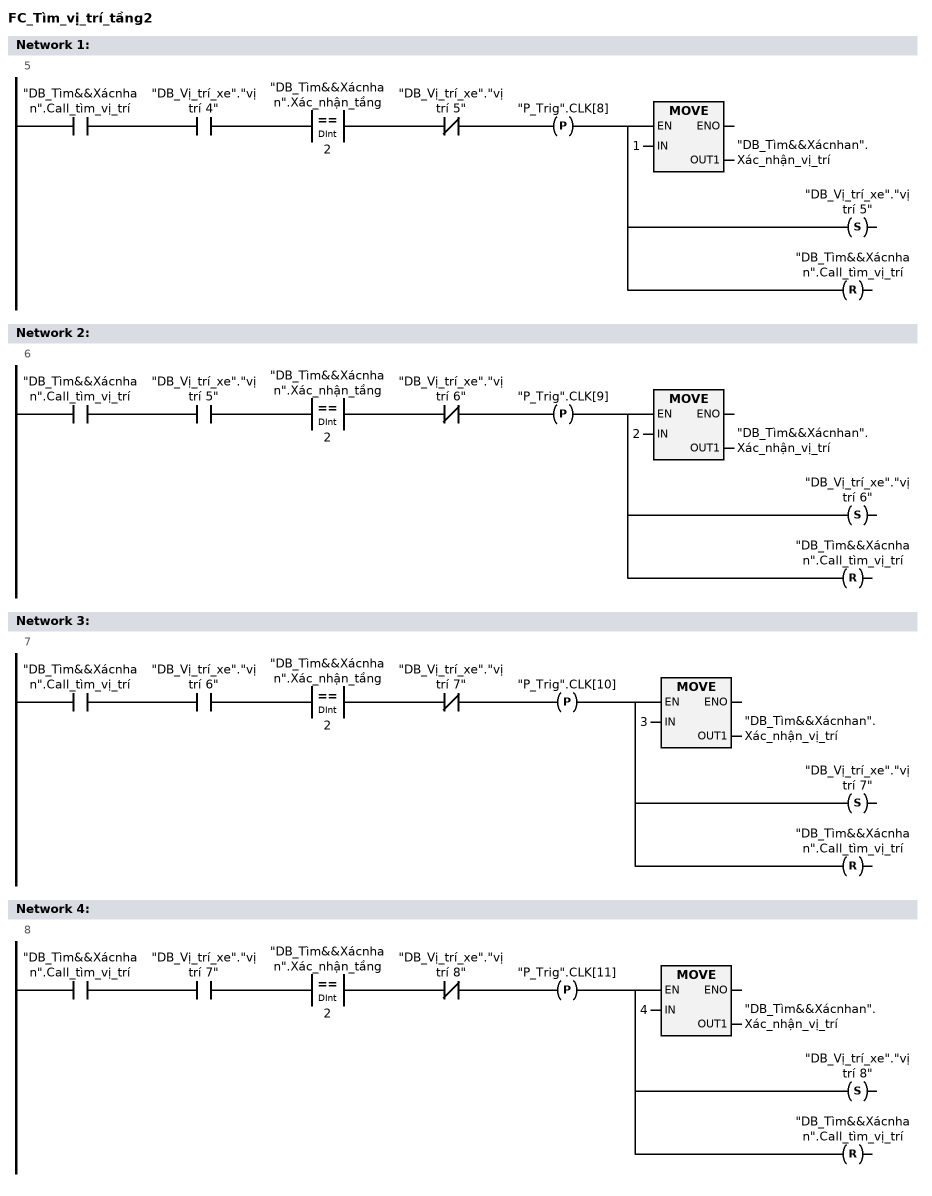
   RUNG wire#powerrail
      Contact( "DB_Tìm&&Xácnhan".Call_tìm_vị_trí )
      Contact( "DB_Vị_trí_xe"."vị trí 4" )
      { S7_Templates := "SrcType := DInt" } EQ_Contact(in1 := "DB_Tìm&&Xácnhan".Xác_nhận_tầng, in2 := 2)
      I_Contact( "DB_Vị_trí_xe"."vị trí 5" )
      P_Trig( "P_Trig".CLK[8] )
      wire#w1
      Move(in := 1, out1 => "DB_Tìm&&Xácnhan".Xác_nhận_vị_trí)
   END_RUNG
   RUNG wire#w1
      S_Coil( "DB_Vị_trí_xe"."vị trí 5" )
   END_RUNG
   RUNG wire#w1
      R_Coil( "DB_Tìm&&Xácnhan".Call_tìm_vị_trí )
   END_RUNG
   // the same network as SCL:
   #_w1 := "DB_Tìm&&Xácnhan".Call_tìm_vị_trí AND "DB_Vị_trí_xe"."vị trí 4" AND ("DB_Tìm&&Xácnhan".Xác_nhận_tầng = 2) AND NOT "DB_Vị_trí_xe"."vị trí 5";
   #_w2 := #_w1 AND NOT "P_Trig".CLK[8];   // rising edge
   "P_Trig".CLK[8] := #_w1;
   IF #_w2 THEN
       "DB_Tìm&&Xácnhan".Xác_nhận_vị_trí := 1;
       "DB_Vị_trí_xe"."vị trí 5" := TRUE;
       "DB_Tìm&&Xácnhan".Call_tìm_vị_trí := FALSE;
   END_IF;
END_REGION

REGION Network 2
   // 6
   RUNG wire#powerrail
      Contact( "DB_Tìm&&Xácnhan".Call_tìm_vị_trí )
      Contact( "DB_Vị_trí_xe"."vị trí 5" )
      { S7_Templates := "SrcType := DInt" } EQ_Contact(in1 := "DB_Tìm&&Xácnhan".Xác_nhận_tầng, in2 := 2)
      I_Contact( "DB_Vị_trí_xe"."vị trí 6" )
      P_Trig( "P_Trig".CLK[9] )
      wire#w1
      Move(in := 2, out1 => "DB_Tìm&&Xácnhan".Xác_nhận_vị_trí)
   END_RUNG
   RUNG wire#w1
      S_Coil( "DB_Vị_trí_xe"."vị trí 6" )
   END_RUNG
   RUNG wire#w1
      R_Coil( "DB_Tìm&&Xácnhan".Call_tìm_vị_trí )
   END_RUNG
   // the same network as SCL:
   #_w1 := "DB_Tìm&&Xácnhan".Call_tìm_vị_trí AND "DB_Vị_trí_xe"."vị trí 5" AND ("DB_Tìm&&Xácnhan".Xác_nhận_tầng = 2) AND NOT "DB_Vị_trí_xe"."vị trí 6";
   #_w2 := #_w1 AND NOT "P_Trig".CLK[9];   // rising edge
   "P_Trig".CLK[9] := #_w1;
   IF #_w2 THEN
       "DB_Tìm&&Xácnhan".Xác_nhận_vị_trí := 2;
       "DB_Vị_trí_xe"."vị trí 6" := TRUE;
       "DB_Tìm&&Xácnhan".Call_tìm_vị_trí := FALSE;
   END_IF;
END_REGION

REGION Network 3
   // 7
   RUNG wire#powerrail
      Contact( "DB_Tìm&&Xácnhan".Call_tìm_vị_trí )
      Contact( "DB_Vị_trí_xe"."vị trí 6" )
      { S7_Templates := "SrcType := DInt" } EQ_Contact(in1 := "DB_Tìm&&Xácnhan".Xác_nhận_tầng, in2 := 2)
      I_Contact( "DB_Vị_trí_xe"."vị trí 7" )
      P_Trig( "P_Trig".CLK[10] )
      wire#w1
      Move(in := 3, out1 => "DB_Tìm&&Xácnhan".Xác_nhận_vị_trí)
   END_RUNG
   RUNG wire#w1
      S_Coil( "DB_Vị_trí_xe"."vị trí 7" )
   END_RUNG
   RUNG wire#w1
      R_Coil( "DB_Tìm&&Xácnhan".Call_tìm_vị_trí )
   END_RUNG
   // the same network as SCL:
   #_w1 := "DB_Tìm&&Xácnhan".Call_tìm_vị_trí AND "DB_Vị_trí_xe"."vị trí 6" AND ("DB_Tìm&&Xácnhan".Xác_nhận_tầng = 2) AND NOT "DB_Vị_trí_xe"."vị trí 7";
   #_w2 := #_w1 AND NOT "P_Trig".CLK[10];   // rising edge
   "P_Trig".CLK[10] := #_w1;
   IF #_w2 THEN
       "DB_Tìm&&Xácnhan".Xác_nhận_vị_trí := 3;
       "DB_Vị_trí_xe"."vị trí 7" := TRUE;
       "DB_Tìm&&Xácnhan".Call_tìm_vị_trí := FALSE;
   END_IF;
END_REGION

REGION Network 4
   // 8
   RUNG wire#powerrail
      Contact( "DB_Tìm&&Xácnhan".Call_tìm_vị_trí )
      Contact( "DB_Vị_trí_xe"."vị trí 7" )
      { S7_Templates := "SrcType := DInt" } EQ_Contact(in1 := "DB_Tìm&&Xácnhan".Xác_nhận_tầng, in2 := 2)
      I_Contact( "DB_Vị_trí_xe"."vị trí 8" )
      P_Trig( "P_Trig".CLK[11] )
      wire#w1
      Move(in := 4, out1 => "DB_Tìm&&Xácnhan".Xác_nhận_vị_trí)
   END_RUNG
   RUNG wire#w1
      S_Coil( "DB_Vị_trí_xe"."vị trí 8" )
   END_RUNG
   RUNG wire#w1
      R_Coil( "DB_Tìm&&Xácnhan".Call_tìm_vị_trí )
   END_RUNG
   // the same network as SCL:
   #_w1 := "DB_Tìm&&Xácnhan".Call_tìm_vị_trí AND "DB_Vị_trí_xe"."vị trí 7" AND ("DB_Tìm&&Xácnhan".Xác_nhận_tầng = 2) AND NOT "DB_Vị_trí_xe"."vị trí 8";
   #_w2 := #_w1 AND NOT "P_Trig".CLK[11];   // rising edge
   "P_Trig".CLK[11] := #_w1;
   IF #_w2 THEN
       "DB_Tìm&&Xácnhan".Xác_nhận_vị_trí := 4;
       "DB_Vị_trí_xe"."vị trí 8" := TRUE;
       "DB_Tìm&&Xácnhan".Call_tìm_vị_trí := FALSE;
   END_IF;
END_REGION
END_FUNCTION

FUNCTION "FC_tìm_vị_trí" : Void   // FC8, LAD
{ S7_Optimized_Access := 'TRUE' }
VERSION : 0.1
BEGIN

REGION Network 1
   // Tìm trong tầng , coi vị trí trống,move hướng(1-4),đánh dấu vị trí,kết thuc gọi tìm vị trí
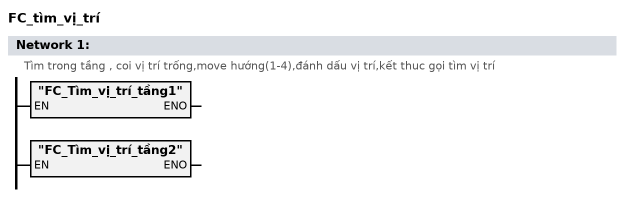
   RUNG wire#powerrail
      "FC_Tìm_vị_trí_tầng1"()
   END_RUNG
   RUNG wire#powerrail
      "FC_Tìm_vị_trí_tầng2"()
   END_RUNG
   // the same network as SCL:
   "FC_Tìm_vị_trí_tầng1"();
   "FC_Tìm_vị_trí_tầng2"();
END_REGION
END_FUNCTION

(* ===== HMI "HMI_RT_1" =====
connection "HMI_Connection_1": ETHERNET, ILRT_S7_1500_OMS

HMI tags "Default tag table"
   "DB_AxisPanel_Lift_Job_Velocity" : Real = PLC DB_AxisPanel.Lift.Job.Velocity, T1s

HMI tags "Operater"
   "DB_Operater_Confirm_Gửi" : Bool = PLC DB_Operater.Confirm_Gửi AT %DB6.DBX0.0, T100ms
   "DB_Operater_Confirm_Lấy" : Bool = PLC DB_Operater.Confirm_Lấy AT %DB6.DBX0.1, T100ms
   "DB_Operater_Scada_Gửi_Xe" : Bool = PLC DB_Operater.Scada_Gửi_Xe AT %DB6.DBX0.3, T100ms
   "DB_Operater_Scada_Lấy_Xe" : Bool = PLC DB_Operater.Scada_Lấy_Xe AT %DB6.DBX0.4, T100ms
   "DB_Operater_ConfirmRFID" : Bool = PLC DB_Operater.ConfirmRFID AT %DB6.DBX0.2, T100ms
   "DB_Operater_Scada_Home_Lift" : Bool = PLC DB_Operater.Scada_Home_Lift AT %DB6.DBX0.6, T100ms
   "DB_Operater_AutoMan" : Bool = PLC DB_Operater.Auto/Man AT %DB6.DBX1.0, T100ms
   "DB_Operater_Static_Mode" : Int = PLC DB_Operater.Static_Mode AT %DB6.DBW2, T100ms

HMI tags "Step"
   "DB_Step_Power" : Bool = PLC DB_Step.Power, T100ms
   "DB_Step_Home_Lift" : Bool = PLC DB_Step.Home.Lift, T100ms
   "DB_Step_Home_Rotation" : Bool = PLC DB_Step.Home.Rotation, T100ms
   "DB_Step_Home_Reach" : Bool = PLC DB_Step.Home.Reach, T100ms
   "DB_Step_HomeAll" : Bool = PLC DB_Step.HomeAll, T100ms
   "DB_Step_ErorrHomeCode_Lift" : Word = PLC DB_Step.ErorrHomeCode.Lift, T100ms
   "DB_Step_ErorrHomeCode_Rotation" : Word = PLC DB_Step.ErorrHomeCode.Rotation, T100ms
   "DB_Step_ErorrHomeCode_Reach" : Word = PLC DB_Step.ErorrHomeCode.Reach, T100ms
   "DB_Step_ErrorHome_Lift" : Bool = PLC DB_Step.ErrorHome.Lift, T100ms
   "DB_Step_ErrorHome_Rotation" : Bool = PLC DB_Step.ErrorHome.Rotation, T100ms
   "DB_Step_ErrorHome_Reach" : Bool = PLC DB_Step.ErrorHome.Reach, T100ms
   "DB_Step_ErorrAbsoluteCode_Rotation" : Word = PLC DB_Step.ErorrAbsoluteCode.Rotation, T100ms
   "DB_Step_ErorrAbsoluteCode_Lift" : Word = PLC DB_Step.ErorrAbsoluteCode.Lift, T100ms
   "DB_Step_ErorrAbsoluteCode_Reach" : Word = PLC DB_Step.ErorrAbsoluteCode.Reach, T100ms
   "DB_Step_ErrorAbsolute_Lift" : Bool = PLC DB_Step.ErrorAbsolute.Lift, T100ms
   "DB_Step_ErrorAbsolute_Rotation" : Bool = PLC DB_Step.ErrorAbsolute.Rotation, T100ms
   "DB_Step_ErrorAbsolute_Reach" : Bool = PLC DB_Step.ErrorAbsolute.Reach, T100ms
   "DB_Step_ErrorJog_Lift" : Word = PLC DB_Step.ErrorJog.Lift, T100ms
   "DB_Step_ErrorJog_Rotation" : Word = PLC DB_Step.ErrorJog.Rotation, T100ms
   "DB_Step_ErrorJog_Reach" : Word = PLC DB_Step.ErrorJog.Reach, T100ms
   "DB_Step_Reset" : Bool = PLC DB_Step.Reset, T100ms
   "DB_Step_PowerStarted" : Bool = PLC DB_Step.PowerStarted, T100ms
   "DB_Step_HomeStarted" : Bool = PLC DB_Step.HomeStarted, T100ms
   "DB_Step_DoneHome" : Bool = PLC DB_Step.DoneHome, T100ms

HMI tags "Convert"
   "DB_Convert_Python_Floor" : Int = PLC DB_Convert.Python.Floor AT %DB14.DBW0, T1s
   "DB_Convert_Python_Location" : Int = PLC DB_Convert.Python.Location AT %DB14.DBW2, T1s
   "DB_Convert_Python_Passcodeplc" : Int = PLC DB_Convert.Python.Passcodeplc AT %DB14.DBW4, T1s
   "DB_Convert_Python_UID" : Array [0..11] of String[14] = PLC DB_Convert.Python.UID AT %DB14.DBX6.0, T1s
   "DB_Convert_Python_Receive" : String[14] = PLC DB_Convert.Python.Receive AT %DB14.DBX198.0, T1s
   "DB_Convert_Floor_Dic1" : Int = PLC DB_Convert.Floor_Dic1 AT %DB14.DBW214, T1s
   "DB_Convert_Floor_Dic2" : Int = PLC DB_Convert.Floor_Dic2 AT %DB14.DBW216, T1s
   "DB_Convert_Location" : Int = PLC DB_Convert.Location AT %DB14.DBW218, T1s
   "DB_Convert_Down" : Int = PLC DB_Convert.Down AT %DB14.DBW220, T1s
   "DB_Convert_Up" : Int = PLC DB_Convert.Up AT %DB14.DBW222, T1s
   "DB_Convert_Started" : Bool = PLC DB_Convert.Started AT %DB14.DBX224.0, T1s

HMI tags "Axis_Panel"
   "DB_AxisPanel_Lift" : UDT = PLC DB_AxisPanel.Lift, T100ms
   "DB_AxisPanel_Rotation" : UDT = PLC DB_AxisPanel.Rotation, T100ms
   "DB_AxisPanel_Reach" : UDT = PLC DB_AxisPanel.Reach, T100ms

HMI tags "Vị trí xe"
   "DB_Vị_trí_xe_vị trí 1" : Bool = PLC DB_Vị_trí_xe."vị trí 1" AT %DB2.DBX0.0, T100ms
   "DB_Vị_trí_xe_vị trí 2" : Bool = PLC DB_Vị_trí_xe."vị trí 2" AT %DB2.DBX0.1, T100ms
   "DB_Vị_trí_xe_vị trí 3" : Bool = PLC DB_Vị_trí_xe."vị trí 3" AT %DB2.DBX0.2, T100ms
   "DB_Vị_trí_xe_vị trí 4" : Bool = PLC DB_Vị_trí_xe."vị trí 4" AT %DB2.DBX0.3, T100ms
   "DB_Vị_trí_xe_vị trí 5" : Bool = PLC DB_Vị_trí_xe."vị trí 5" AT %DB2.DBX0.4, T100ms
   "DB_Vị_trí_xe_vị trí 6" : Bool = PLC DB_Vị_trí_xe."vị trí 6" AT %DB2.DBX0.5, T100ms
   "DB_Vị_trí_xe_vị trí 7" : Bool = PLC DB_Vị_trí_xe."vị trí 7" AT %DB2.DBX0.6, T100ms
   "DB_Vị_trí_xe_vị trí 8" : Bool = PLC DB_Vị_trí_xe."vị trí 8" AT %DB2.DBX0.7, T100ms
   "DB_Vị_trí_xe_tầng_1" : Bool = PLC DB_Vị_trí_xe.tầng_1 AT %DB2.DBX1.0, T100ms
   "DB_Vị_trí_xe_tầng_2" : Bool = PLC DB_Vị_trí_xe.tầng_2 AT %DB2.DBX1.1, T100ms

text list "SystemTextList_ConfigErrorAlarmTextLibrary_1": 1 'NameService configuration error: Implicit deletion. Subelement instance @6%s@ must be deleted explicitly.'; 2 'NameService configuration error: Implicit deletion. Alias/Format/Unit instance @6%s@ must be deleted explicitly.'

text list "SystemTextList_ConfigErrorAlarmTextLibrary_2": 1 'EvDpManager::cleanupDeletedDatapoint - alert handler config is deleted implicitly for deleted datapoint, @3%s@'; 2 'EvDpManager::cleanupDeletedDatapoint - alert handler config is deleted implicitly but still has overrides, @3%s@'; 3 'EvDpManager::cleanupDeletedDatapoint - default value config is deleted implicitly for deleted datapoint, @3%s@'; 4 'EvDpManager::cleanupDeletedDatapoint - default value config is deleted implicitly but still has overrides, @3%s@'; 5 'EvDpManager::cleanupDeletedDatapoint - initial value config is deleted implicitly for deleted datapoint, @3%s@'; 6 'EvDpManager::cleanupDeletedDatapoint - initial value config is deleted implicitly but still has overrides, @3%s@'; 7 'EvDpManager::cleanupDeletedDatapoint - distribution config is deleted implicitly for deleted datapoint, @3%s@'; 8 'EvDpManager::cleanupDeletedDatapoint - distribution config is deleted implicitly but still has overrides, @3%s@'; 9 'EvDpManager::cleanupDeletedDatapoint - rangeCheck config is deleted implicitly for deleted datapoint, @3%s@'; 10 'EvDpManager::cleanupDeletedDatapoint - rangeCheck config is deleted implicitly but still has overrides, @3%s@'

text list "SystemTextList_ConfigErrorAlarmTextLibrary_3": 1 'The configured data point type was deleted, but a configured type is still defined for the node type: @3%s@.'; 2 'The configured data point node type was deleted in the data point type, but a configured type is still defined for the element: @3%s@.'

text list "SystemTextList_ConfigErrorAlarmTextLibrary_4": 2 'Cycles: @6%s@ does not exist'; 3 'Alarms: @6%s@ exists already'; 4 'Tags: Address @6%s@ was rejected'; 1 'Connections: @6%s@ does not exist'; 5 'Tags: Acquisition mode @6%s@ is not supported.'; 6 'Cycles: @6%s@ was deleted but associated tags exist.'; 7 'Connections: @6%s@ was deleted but associated tags exist.'; 8 'Tags: Tag @6%s@ was rejected.'; 9 'Tags: Tag @6%s@ has an invalid value.'; 0 'Connections: Connection to @6%s@ could not be established.'; 65638 'Connections: Connection to @6%s@ could not be established.'; 65639 'Connections: @6%s@ disconnected.'; 65640 'Connections: Connection to the HMI device @6%s@ is lost.'; 65641 'Connections: Connection to the PLC @6%s@ is lost.'; 65541 'Connections: Timeout while establishing the connection to @6%s@.'; 65542 'Connections: @6%s@ faulty.'; 65543 'Connections: Connection to the HMI device disconnected. Connection @5%s@ was changed.'; 65544 'Connections: Connection to the HMI device disconnected. Driver property was changed for connection @5%s@.'

text list "SystemTextList_ConfigErrorAlarmTextLibrary_5": 1 'Connections: Lifecycle monitoring cycle must be shorter than the response time.'; 2 'Connections: Cyclic services are configured but not supported by the target device.'; 3 'Connections: Change-controlled reading is configured but not supported by the target device.'; 4 'Tags: The address @6%s@ does not exist in the PLC.'; 5 'Tags: The default conversion type for the address @6%s@ could not be determined.'; 6 'Tags: Invalid conversion type'; 7 'Cycles: Invalid conversion type. Conversion is not supported at HmiCycle.'; 4096 'Connections: Version of the address @6%s@ is not supported.'; 4097 'Connections: PROFIBUS address is not supported.'; 4098 'Connections: Softbus address is not supported.'; 4099 'Connections: Address type @6%s@ is not supported.'; 4100 'Connections: Invalid connection name @6%s@. Access point is being ignored.'; 4101 'Connections: Routing is not supported. @6%s@ is not used.'; 4102 'Connections: Routing is not supported. @6%s@ is not used.'; 4103 'Connections: Invalid IP address @6%s@'; 4104 'Connections: Invalid Named Connection @6%s@. Valid format: >VMD</>connection<'; 4105 'Connections: Invalid Named Connection @6%s@. VMD connection name is too long. Only 24 characters are permitted.'; 4106 'Connections: Invalid Named Connection @6%s@. Connection name is too long. Only 32 characters are permitted.'; 4107 'Connections: Rack number @6%s@ is outside of the permitted range (0..7)'; 4108 'Connections: Invalid Named Connection @6%s@. Rack is ignored.'; 4109 'Connections: Slot number @6%s@ is outside of the permitted range (1..32)'; 4110 'Connections: Invalid Named Connection @6%s@. Slot is ignored.'; 4111 'Connection could not be established. Maximum number of available connections (@6%s@) has been exceeded.'; 4112 'Connection aborted. No sign of life in the last @4%s@ ms.'; 4113 'Connection could not be established - @4%s@'; 4114 'Connection could not be established. The address @6%s@ cannot be used.'; 4115 'Connection could not be established. Invalid address @6%s@'; 4116 'Connection could not be established - @4%s@'

text list "SystemTextList_ConfigErrorAlarmTextLibrary_6": 1 'Connection could not be established. Application instance certificate is not configured.'; 2 'Connection could not be established. Server has rejected the client certificate. OPC UA status code @4%s@.'; 3 'Connection could not be established. Internal problem in the certificate store. OPC UA status code @4%s@'; 4 'Connection could not be established. Application instance certificate could not be loaded. OPC UA status code @4%s@'; 5 'Connection could not be established. Server has not provided a certificate. @4%s@'; 6 'Connection could not be established. Validation of server certificate has failed. OPC UA status code @4%s@.'; 7 'Connection was closed. Error during alarm synchronization. OPC UA status code @4%s@.'; 8 'Connection was closed. Alarm/event subscription has failed. The number of operations on the server has been exceeded.'; 9 'Connection was closed. Alarm/event subscription has failed. The number of alarm/event subscriptions on the server has been exceeded.'; 10 'Connection could not be established. Server reports a license problem. OPC UA status code @4%s@.'; 11 'Connection could not be established. Maximum number of server sessions has been exceeded.'; 12 'Connection could not be established. Safety configuration is inconsistent. @4%s@'; 13 'Connection could not be established. The address @4%s@ cannot be used.'; 14 'Connection could not be established. OPC UA status code @4%s@'; 15 'Connection aborted. OPC UA server was stopped.'; 16 'Connection aborted. No sign of life in the last @4%s@ ms.'; 17 'Connection was closed. OPC UA server maintenance.'; 18 'Connection could not be established. Invalid configuration of the authentication mode - @4%s@'; 19 'Connection could not be established. User could not be authenticated. OPC UA status code @4%s@'; 20 'Connection could not be established. Server does not permit anonymous connection. OPC UA status code @4%s@'; 21 'Connection could not be established. Certificate problem: Error when writing the safety-relevant data to @4%s@.'; 22 'Connection could not be established. Certificate problem: Unexpected file in the folder @4%s@ cannot be removed.'; 23 'Connection could not be established. User could not be authenticated. No user or password configured.'; 24 'Connection could not be established. Unexpected length of the server certificate. @4%s@'; 25 'Connection could not be established. @4%s@ is empty.'; 26 'Connection could not be established. @4%s@ has an unexpected format.'; 27 'Connection could not be established. Server endpoints cannot be read. OPC UA status code @4%s@'; 28 'Connection could not be established. No server endpoints were found. @4%s@'; 29 'Connection could not be established. Application instance certificate could not be found.'; 30 'Connection could not be established. Unexpected format of the certificate @4%s@.'; 31 'Connection could not be established. Unexpected format of the certificate block list @4%s@.'; 32 'Connection could not be established. User could not be authenticated. An encryption detail is invalid. @4%s@'; 34 'Connection could not be established. - The configured non-transparent redundancy mode @4%s@ is not supported.'; 101 'Tags: Address @6%s@ does not exist on the server.'; 103 'Tags: Address @6%s@ cannot be accessed.'; 104 'Tags: Acquisition mode is not supported for address @6%s@.'; 201 'Alarms: Address @6%s@ does not exist on the server.'; 202 'Alarms: Address @6%s@ cannot be used. The specified range filter is not an OPC UA Event Notifier.'; 203 'Alarms: Address @6%s@ cannot be used. The specified range filter does not exist on the server.'; 204 'Alarms: Address @6%s@ cannot be used because it is not an OPC UA event type.'; 205 'Alarms: Address @6%s@ cannot be used because the OPC UA condition type is not supported.'; 206 'Alarms: Address @6%s@ cannot be used because the event type does not exist on the server.'; 207 'Alarms: Acquisition type cannot be used for address @6%s@.'; 301 'Address @6%s@ cannot be used because the version number is missing.'; 302 'Address @6%s@ cannot be used because the version number is invalid.'; 303 'Address @6%s@ cannot be used because the number of '$' delimiters is invalid.'; 304 'Address @6%s@ cannot be used because the address type is invalid.'; 305 'Unsupported version @6%s@ of the address'; 401 'Unexpected OPC UA server response: @6%s@'

text list "SystemTextList_ConfigErrorAlarmTextLibrary_7": 1 'Messages: Invalid condition string for the alarm view @6%s@.'; 2 'Messages: Invalid status tag and bit for the alarm view @6%s@.'; 3 'Messages: Invalid control tag and bit for the alarm view @6%s@.'

text list "SystemTextList_ConfigErrorAlarmTextLibrary_8": 1 'Logs: Implicit deletion. Logging tag instance @6%s@ should be deleted but there are overloaded elements.'

text list "SystemTextList_ConfigErrorAlarmTextLibrary_9": 1 ''; 2 'Restart of the runtime is required.'; 3 'The correct storage medium must be ejected and inserted again.'

text list "SystemTextList_ConfigErrorAlarmTextLibrary_10": 1 'CDS cache - Cache folder cannot be created or reached: @6%s@'; 2 'LOC cache - Cache folder cannot be created or reached: @6%s@'

text list "SystemTextList_RuntimeCollaborationFailureReason_1": 0 'Unknown error (@3%s@)'; 1 'The system is not running or there is a network problem'; 2 'Runtime is not started on the target device.'; 3 'The System ID does not match the expected System ID (@3%s@)'; 4 'The Collaboration name does not match the expected Collaboration name '@3%s@''; 5 'Wrong or unknown certificate'; 6 'Revoked certificate'; 7 'The time difference is too big.'; 8 'No common supported message version'; 9 'System ID (@3%s@) already exists'; 10 'System name (@3%s@) already exists'; 11 'ID/Name in local configuration for Runtime Collaboration already exists'

text list "SystemTextList_S7PlusAlarmTextListCollection_1": 4096 'Connections: Connection to the PLC @4%s@ is lost'; 4097 'Connections: Connection to the HMI device @4%s@ is lost'; 4098 'Connections: Maximum number of connections exceeded - @4%s@'; 4099 'Out of resources on PLC - @4%s@'; 4100 'Legitimation failed, invalid or missing password - @4%s@'; 4101 'Request to open the connection failed - @4%s@'; 4102 'Connections: Cannot connect to PLC - @4%s@'; 4103 'Request to open the connection could not be sent'; 4104 'General certificate error for PLC - @4%s@'; 4105 'PLC certificate expired for PLC - @4%s@'; 4106 'PLC certificate is revoked for PLC - @4%s@'; 4107 'PLC certificate is untrustworthy. Manual trust is possible for - @4%s@'; 4108 'PLC certificate is untrustworthy. Manual trust is not possible for - @4%s@'

text list "SystemTextList_AllenBradleyEIPAlarmTextListCollection_7": 4096 'Connection lost on PLC side - @5%s@'; 4097 'Connection lost on HMI side - @5%s@'; 4098 'Maximum number of connections exceeded - @5%s@'; 4099 'Out of resources on PLC - @5%s@'; 4100 'Legitimation failed, invalid or missing password - @5%s@'; 4101 'Open request failed - @5%s@'; 4102 'Cannot connect to PLC - @5%s@'; 4103 'Open request could not be sent'; 4104 'root certificate expired for - @5%s@'; 4105 'PLC certificate untrusted for - @5%s@'

text list "SystemTextList_OmronEIPAlarmTextListCollection_6": 4096 'Connection lost on PLC side - @5%s@'; 4097 'Connection lost on HMI side - @5%s@'; 4098 'Maximum number of connections exceeded - @5%s@'; 4099 'Out of resources on PLC - @5%s@'; 4100 'Legitimation failed, invalid or missing password - @5%s@'; 4101 'Open request failed - @5%s@'; 4102 'Cannot connect to PLC - @5%s@'; 4103 'Open request could not be sent'; 4104 'root certificate expired for - @5%s@'; 4105 'PLC certificate untrusted for - @5%s@'

text list "SystemTextList_StdModbusTCPAlarmTextListCollection_5": 4096 'Connections: Connection to the PLC @5%s@ is lost'; 4097 'Connections: Connection to the HMI device @5%s@ is lost'; 4098 'Connections: Maximum number of connections exceeded - @5%s@'; 4099 'Out of resources on PLC - @5%s@'; 4100 'Legitimation failed, invalid or missing password - @5%s@'; 4101 'Request to open the connection failed - @5%s@'; 4102 'Connections: Cannot connect to PLC - @5%s@'; 4103 'Request to open the connection could not be sent'; 4104 'General certificate error for PLC - @5%s@'; 4105 'PLC certificate expired for PLC - @5%s@'; 4106 'PLC certificate is revoked for PLC - @5%s@'; 4107 'PLC certificate is untrustworthy. Manual trust is possible for - @5%s@'; 4108 'PLC certificate is untrustworthy. Manual trust is not possible for - @5%s@'

text list "SystemTextList_MitsubishiMCAlarmTextListCollection_4": 4096 'Connection lost on PLC side - @5%s@'; 4097 'Connection lost on HMI side - @5%s@'; 4098 'Maximum number of connections exceeded - @5%s@'; 4099 'Out of resources on PLC - @5%s@'; 4100 'Legitimation failed, invalid or missing password - @5%s@'; 4101 'Open request failed - @5%s@'; 4102 'Cannot connect to PLC - @5%s@'; 4103 'Open request could not be sent'; 4104 'root certificate expired for - @5%s@'; 4105 'PLC certificate untrusted for - @5%s@'

text list "SystemTextList_MitsubishiiQAlarmTextListCollection_3": 4096 'Connection lost on PLC side - @5%s@'; 4097 'Connection lost on HMI side - @5%s@'; 4098 'Maximum number of connections exceeded - @5%s@'; 4099 'Out of resources on PLC - @5%s@'; 4100 'Legitimation failed, invalid or missing password - @5%s@'; 4101 'Open request failed - @5%s@'; 4102 'Cannot connect to PLC - @5%s@'; 4103 'Open request could not be sent'; 4104 'root certificate expired for - @5%s@'; 4105 'PLC certificate untrusted for - @5%s@'

text list "SystemTextList_StdModbusRTUAlarmTextListCollection_8": 4096 'Connections: Connection to the PLC @5%s@ is lost'; 4097 'Connections: Connection to the HMI device @5%s@ is lost'; 4098 'Connections: Maximum number of connections exceeded - @5%s@'; 4099 'Out of resources on PLC - @5%s@'; 4100 'Legitimation failed, invalid or missing password - @5%s@'; 4101 'Request to open the connection failed - @5%s@'; 4102 'Connections: Cannot connect to PLC - @5%s@'; 4103 'Request to open the connection could not be sent'; 4104 'General certificate error for PLC - @5%s@'; 4105 'PLC certificate expired for PLC - @5%s@'; 4106 'PLC certificate is revoked for PLC - @5%s@'; 4107 'PLC certificate is untrustworthy. Manual trust is possible for - @5%s@'; 4108 'PLC certificate is untrustworthy. Manual trust is not possible for - @5%s@'

text list "Static_Mode": -1 ''; 1 'AUTO'; 2 'MANUAL'
*)

(* ===== HMI "HiddenHmiRTDeviceFaceplateTypes" =====

HMI tags "8f57ea34-786a-4f61-8df0-d11cb035e70c"
   "Tiltle" : WString[254], internal
*)

(* ===== HMI "HiddenHmiRTDeviceFaceplateTypes" =====

HMI tags "8f57ea34-786a-4f61-8df0-d11cb035e70c"
   "Tiltle" : WString[254], internal
*)

(* ===== HMI "HiddenHmiRTDeviceFaceplateTypes" =====

HMI tags "8f57ea34-786a-4f61-8df0-d11cb035e70c"
   "Tiltle" : WString[254], internal
*)